// Mitsubishi GX Works2 project: 化成1_Debug 5.21   PLC: Q06UDEH

TYPE SwitchIO : STRUCT
  xLiftCylinderRetractDetect : BOOL;
  xLiftCylinderExtendDetect : BOOL;
  xLiftCylinderRetract : BOOL;
  xLiftCylinderExtend : BOOL;
  xEntryBarCylinderRetract : BOOL;
  xLiftCylinderExtendInit : BOOL;
  xEntryEnable : BOOL;
  xExitEnable : BOOL;
  xExitBarCylinderRetract : BOOL;
  xSwithEnable : BOOL;
  xLiftCylinderRetractButton : BOOL;
  xLiftCylinderExtendButton : BOOL;
  xEntryBarCylinderRetractButton : BOOL;
  xExitBarCylinderRetractButton : BOOL;
END_STRUCT END_TYPE

TYPE ConveyorIO : STRUCT
  iProductCategory : INT;  (* 产品类型0：无料1：正极  2：负极 3：隔膜 4：空料架 *)
  xCWPresent : BOOL;  (* 正转检测有无传感器 *)
  xCCWPresent : BOOL;  (* 反转检测有无传感器 *)
  xLoad : BOOL;  (* 上料请求 *)
  xUnload : BOOL;  (* 下料请求 *)
  xMotorCW : BOOL;  (* 电机正转 *)
  xMotorCCW : BOOL;  (* 电机反转 *)
  xEmpty : BOOL;  (* 线体状态为空 *)
  xNextRun : BOOL;  (* 下段线体运行 *)
  xUnloadCCW : BOOL;  (* 下料为反转 *)
  xloadCCW : BOOL;  (* 上料为反转 *)
  xLeave : BOOL;  (* 已经离开 *)
  xForward : BOOL;  (* 正转手动 *)
  xBackward : BOOL;  (* 反转手动 *)
  xBusy : BOOL;  (* 工作中 *)
  tLoadDelay : TIME;  (* 进入延时设置 *)
  xPutInto : BOOL;  (* 线体直接投入物料 *)
  xUnloadAlarm : BOOL;  (* 下料报警 *)
  xPosLimit : BOOL;  (* 正限位 *)
  xNegLimit : BOOL;  (* 负限位 *)
  xOverWidthAlarm : BOOL;  (* 超宽报警 *)
  xLimitAlarrm : BOOL;  (* 限位报警 *)
  iDeviceID : INT;  (* 线体ID *)
  xSizeDeficientDetect : BOOL;  (* 尺寸不足检测标志位 *)
END_STRUCT END_TYPE

TYPE ShuttleCarIO : STRUCT
  xReady : BOOL;  (* 准备就绪 *)
  xForward : BOOL;  (* 正转 *)
  xBackward : BOOL;  (* 反转 *)
  iCurrentPos : INT;  (* 当前位置 *)
  iDestinationPos : INT;  (* 目标位置 *)
  xCW : BOOL;  (* 正转输出 *)
  xCCW : BOOL;  (* 反转输出 *)
  xBrake : BOOL;  (* 刹车 *)
  xHomeSwitch : BOOL;  (* 零位接近开关 *)
  xPosLimit : BOOL;  (* 正限位 *)
  xNegLimit : BOOL;  (* 负限位 *)
  xMDIExe : BOOL;  (* MDI开始 *)
  xMDIDone : BOOL;  (* MDI 完成 *)
  xPassLimit : BOOL;  (* 限位屏蔽 *)
  xPosLimitCatch : BOOL;  (* 正限位捕捉 *)
  xNegLimitCatch : BOOL;  (* 负限位捕捉 *)
  xHomeExe : BOOL;  (* 开始寻零 *)
  xHomeDone : BOOL;  (* 寻零完成 *)
  xHomeBusy : BOOL;  (* 寻零中 *)
  xHomeFailed : BOOL;  (* 寻零失败 *)
  xBusy : BOOL;  (* 工作中 *)
  tArriveDelay : TIME;  (* 到位延时 *)
  xCylinder : BOOL;  (* 气缸控制 *)
  tBrakeDelay : TIME;  (* 抱闸延时 *)
  xPauseRamp : BOOL;  (* 暂停减速斜坡标志位 *)
  xPresentDetect1 : BOOL;  (* 物料有无检测1 *)
  xPresentDetect2 : BOOL;  (* 物料有无检测2 *)
  xOvertimeAlarm : BOOL;  (* 超时报警 *)
  tSetOverTime : TIME;  (* 设置超时时间 *)
  xLooseDetect : BOOL;  (* 松绳检测 *)
  xLooseAlarm : BOOL;  (* 松绳报警 *)
END_STRUCT END_TYPE

TYPE Stub : STRUCT
  xLoadRequest : BOOL;
  xLoadRequestAkn : BOOL;
  xUnloadRequest : BOOL;
  xUnloadRequestAkn : BOOL;
END_STRUCT END_TYPE

TYPE RGVCommunication : STRUCT
  xFullLoadRequest : BOOL;  (* 满框上料请求 *)
  xFullUnloadRequest : BOOL;  (* 满框下料请求 *)
  xEmptyLoadRequest : BOOL;  (* 空框上料请求 *)
  xEmptyUnloadRequest : BOOL;  (* 空框下料请求 *)
  xFullLoadRequestAkn : BOOL;  (* 满框上料请求确认 *)
  xFullUnloadRequestAkn : BOOL;  (* 满框下料请求确认 *)
  xEmptyLoadRequestAkn : BOOL;  (* 空框上料请求确认 *)
  xEmptyUnloadRequestAkn : BOOL;  (* 空框下料请求确认 *)
  xFullLoadComplete : BOOL;  (* 满框上料完成 *)
  xFullUnloadComplete : BOOL;  (* 满框下料完成 *)
  xEmptyLoadComplete : BOOL;  (* 空框上料完成 *)
  xEmptyUnloadComplete : BOOL;  (* 空框下料完成 *)
  xFullLoadCompleteAkn : BOOL;  (* 满框上料完成确认 *)
  xFullUnloadCompleteAkn : BOOL;  (* 满框下料完成确认 *)
  xEmptyLoadCompleteAkn : BOOL;  (* 空框上料完成确认 *)
  xEmptyUnloadCompleteAkn : BOOL;  (* 空框下料完成确认 *)
  xMdiExe : BOOL;  (* RGV 执行 *)
  xMdiDone : BOOL;  (* RGV 执行完成 *)
  iCurrentPostion : INT;  (* RGV当前位置 *)
  iDestinationPos : INT;  (* RGV目标位置 *)
  xEmpty1 : BOOL;
  xNextRun1 : BOOL;
  xEmpty2 : BOOL;
  xNextRun2 : BOOL;
  xLoad1 : BOOL;
  xUnload1 : BOOL;
  xLoad2 : BOOL;
  xUnload2 : BOOL;
  xCollisionAlarm : BOOL;  (* 干涉报警 *)
  xRemoteReset : BOOL;  (* 远程复位 *)
  xAuto : BOOL;  (* 自动 *)
END_STRUCT END_TYPE

TYPE BarCylinderIO : STRUCT
  xPresentSwitch : BOOL;  (* 行程开关 *)
  xBarCylinder : BOOL;  (* 阻挡气缸 *)
  xEmpty : BOOL;  (* 为空指示 *)
  xTransportMotorCW : BOOL;  (* 输送电机正转 *)
  xUnload : BOOL;  (* 下料 *)
  xBarCylinderButton : BOOL;  (* 阻挡气缸 *)
  xTransportMotorCWButton : BOOL;  (* 输送电机正转按钮 *)
  xLoad : BOOL;  (* 上料 *)
  xNextRun : BOOL;  (* 下位设备开始运行 *)
  xTransportMotorCCWButton : BOOL;  (* 输送电机反转按钮 *)
  xTransportMotorCCW : BOOL;  (* 输送电机反转 *)
  iProductCategory : INT;  (* 产品种类 *)
  tLoadDelay : TIME;  (* 上料延时 *)
  xBarCylinderSecondary : BOOL;  (* 阻挡第二个无料的气缸 *)
  xBarSecondaryButton : BOOL;  (* 阻挡第二个无料的气缸手动按钮 *)
  iDeviceID : INT;  (* 设备编号 *)
END_STRUCT END_TYPE

// global labels: Global1
VAR_GLOBAL
  g_xAuto AT M11 : BOOL;
  g_xManual : BOOL;
  g_xEStop AT X23 : BOOL;
  g_xReset AT X20 : BOOL;
  g_xStackLampRed AT Y120 : BOOL;
  g_xStackLampAmber AT Y121 : BOOL;
  g_xStackLampGreen AT Y122 : BOOL;
  g_xBuzzer AT Y123 : BOOL;
  g_xStop AT M2 : BOOL;
  g_xLocalAutoStart AT M1 : BOOL;
  g_xRemoteAutoStart AT M0 : BOOL;
  g_xRemoteAuto AT M10 : BOOL;
  g_iState AT D40 : INT;
  g_iLocalAutoStep : BOOL;
  g_xAlarm : BOOL;
  g_xImport1Forbidden AT M174 : BOOL;  (* 1表示禁止从注液入库 *)
  g_xExportChemForbidden AT M176 : BOOL;  (* 1表示禁止出库到化成 *)
  g_xExportBackForbidden AT M177 : BOOL;  (* 1表示禁止返回注液 *)
  g_xImport2Forbidden AT M175 : BOOL;  (* 1表示禁止从化成入库 *)
  g_xResetSingle AT M4 : BOOL;  (* 单线体复位 *)
  g_xInsertTask AT M5 : BOOL;  (* 插入任务 *)
  g_iInsertTask AT D2 : INT;  (* 插入任务号 *)
  g_xPause AT M3 : BOOL;  (* 暂停 *)
  g_iDeviceIDSelect AT D0 : INT;
END_VAR

// global labels: Global
VAR_GLOBAL
  g_xChem2ComFailed : BOOL;
  g_xFillingRGVComFailed : BOOL;
END_VAR

// task Task_01 (event TRUE, interval 0, priority 31): POU, Start, UDP

PROGRAM POU
VAR
  H3000Conveyor1 : Conveyor;
  H3000Conveyor1IO : ConveyorIO;
  H3000Conveyor2 : Conveyor;
  H3000Conveyor2IO : ConveyorIO;
  H3000Conveyor3 : Conveyor;
  H3000Conveyor3IO : ConveyorIO;
  H3000Conveyor4 : Conveyor;
  H3000Conveyor4IO : ConveyorIO;
  H3000Conveyor5 : Conveyor;
  H3000Conveyor5IO : ConveyorIO;
  H3000Conveyor6 : Conveyor;
  H3000Conveyor6IO : ConveyorIO;
  H3000Conveyor7 : Conveyor;
  H3000Conveyor7IO : ConveyorIO;
  H3000Conveyor8 : Conveyor;
  H3000Conveyor8IO : ConveyorIO;
  H3000Conveyor9 : Conveyor;
  H3000Conveyor9IO : ConveyorIO;
  H3000Conveyor10 : Conveyor;
  H3000Conveyor10IO : ConveyorIO;
  H3000ChemConveyor1 : Conveyor;
  H3000ChemConveyor1IO : ConveyorIO;
  H3000ChemConveyor2 : Conveyor;
  H3000ChemConveyor2IO : ConveyorIO;
  H3000ChemConveyor3 : Conveyor;
  H3000ChemConveyor3IO : ConveyorIO;
  Lifter1 : ShuttleCar;
  Lifter1IO : ShuttleCarIO;
  Conveyor1 : Conveyor;
  Conveyor1IO : ConveyorIO;
  Lifter2 : ShuttleCar;
  Lifter2IO : ShuttleCarIO;
  Conveyor2 : Conveyor;
  Conveyor2IO : ConveyorIO;
  H2200Conveyor1 : Conveyor;
  H2200Conveyor1IO : ConveyorIO;
  H2200Conveyor2 : Conveyor;
  H2200Conveyor2IO : ConveyorIO;
  H2200Conveyor3 : Conveyor;
  H2200Conveyor3IO : ConveyorIO;
  H2200Conveyor4 : Conveyor;
  H2200Conveyor4IO : ConveyorIO;
  H2200Conveyor5 : Conveyor;
  H2200Conveyor5IO : ConveyorIO;
  H2200Conveyor6 : Conveyor;
  H2200Conveyor6IO : ConveyorIO;
  H2200Conveyor7 : Conveyor;
  H2200Conveyor7IO : ConveyorIO;
  H2200Conveyor8 : Conveyor;
  H2200Conveyor8IO : ConveyorIO;
  H2200Conveyor9 : Conveyor;
  H2200Conveyor9IO : ConveyorIO;
  H2200Conveyor10 : Conveyor;
  H2200Conveyor10IO : ConveyorIO;
  H1000Conveyor1 : Conveyor;
  H1000Conveyor1IO : ConveyorIO;
  H1000Conveyor2 : Conveyor;
  H1000Conveyor2IO : ConveyorIO;
  H1000Conveyor3 : Conveyor;
  H1000Conveyor3IO : ConveyorIO;
  H1000Conveyor4 : Conveyor;
  H1000Conveyor4IO : ConveyorIO;
  H1000Conveyor5 : Conveyor;
  H1000Conveyor5IO : ConveyorIO;
  H1000Conveyor6 : Conveyor;
  H1000Conveyor6IO : ConveyorIO;
  H1000Conveyor7 : Conveyor;
  H1000Conveyor7IO : ConveyorIO;
  H1000Conveyor8 : Conveyor;
  H1000Conveyor8IO : ConveyorIO;
  H1000Conveyor9 : Conveyor;
  H1000Conveyor9IO : ConveyorIO;
  H3000SwitchChem : Switch;
  H3000SwitchChemIO : SwitchIO;
  H850Switch : Switch;
  H850SwitchIO : SwitchIO;
  H850SwitchConveyorIn : ConveyorIO;
  H850SwitchConveyorOut : ConveyorIO;
  H850Conveyor8 : Conveyor;
  H850Conveyor8IO : ConveyorIO;
  H1000Conveyor10 : Conveyor;
  H1000Conveyor10IO : ConveyorIO;
  H3000SwitchChemConveyorIn : ConveyorIO;
  H3000SwitchChemConveyorOut : ConveyorIO;
  H3000SwitchQuadPackage : Switch;
  H3000SwitchQuadPackageIO : SwitchIO;
  H3000SwitchPackageConveyorIn : ConveyorIO;
  H3000SwitchPackageConveyorOut : ConveyorIO;
  H2200Switch1 : Switch;
  H2200Switch1IO : SwitchIO;
  H2200Switch1ConveyorIn : ConveyorIO;
  H2200Switch1ConveyorOut : ConveyorIO;
  H2200Switch2 : Switch;
  H2200Switch2IO : SwitchIO;
  H2200Switch2ConveyorIn : ConveyorIO;
  H2200Switch2ConveyorOut : ConveyorIO;
  iStep : INT;
  Import1Conveyor1 : Conveyor;
  Import1Conveyor1IO : ConveyorIO;
  Import1Conveyor2 : Conveyor;
  Import1Conveyor2IO : ConveyorIO;
  Import2Conveyor1 : Conveyor;
  Import2Conveyor1IO : ConveyorIO;
  Import2Conveyor2 : Conveyor;
  Import2Conveyor2IO : ConveyorIO;
  Export1Conveyor1 : Conveyor;
  Export1Conveyor1IO : ConveyorIO;
  Export1Conveyor2 : Conveyor;
  Export1Conveyor2IO : ConveyorIO;
  Export2Conveyor1 : Conveyor;
  Export2Conveyor1IO : ConveyorIO;
  Export2Conveyor2 : Conveyor;
  Export2Conveyor2IO : ConveyorIO;
  Export2Switch : Switch;
  Export2SwitchIO : SwitchIO;
  Export2SwitchConveyorIn : ConveyorIO;
  Export2SwitchConveyorOut : ConveyorIO;
  H850Rotor : ShuttleCar;
  H850RotorIO : ShuttleCarIO;
  H850RotorConveyor : Conveyor;
  H850RotorConveyorIO : ConveyorIO;
  H2200RotorIO : ShuttleCarIO;
  H2200RotorConveyor : Conveyor;
  H2200RotorConveyorIO : ConveyorIO;
  H2200Rotor : ShuttleCar;
  H850Conveyor1 : Conveyor;
  H850Conveyor1IO : ConveyorIO;
  H850Conveyor3 : Conveyor;
  H850Conveyor3IO : ConveyorIO;
  H850Conveyor4 : Conveyor;
  H850Conveyor4IO : ConveyorIO;
  H850Conveyor5 : Conveyor;
  H850Conveyor5IO : ConveyorIO;
  H850Conveyor6 : Conveyor;
  H850Conveyor6IO : ConveyorIO;
  Lifter2Position : ARRAY [0..5] OF INT;
  ii : INT;  (* 提升机2任务号 *)
  H2200SwitchEmptyABack : Switch;
  H2200SwitchEmptyABackIO : SwitchIO;
  H2200SwitchEmptyABackConveyorIn : ConveyorIO;
  H2200SwitchEmptyABackConveyorOut : ConveyorIO;
  H2200SwitchEmptyBBack : Switch;
  H2200SwitchEmptyBBackIO : SwitchIO;
  H2200SwitchEmptyBBackConveyorIn : ConveyorIO;
  H2200SwitchEmptyBBackConveyorOut : ConveyorIO;
  H2200ImportConveyor1 : Conveyor;
  H2200ImportConveyor1IO : ConveyorIO;
  H2200ImportConveyor2 : Conveyor;
  H2200ImportConveyor2IO : ConveyorIO;
  Import1Switch : Switch;
  Import1SwitchIO : SwitchIO;
  Import1SwitchConveyorIn : ConveyorIO;
  Import1SwitchConveyorOut : ConveyorIO;
  Export1Switch : Switch;
  Export1SwitchIO : SwitchIO;
  Export1SwitchConveyorIn : ConveyorIO;
  Export1SwitchConveyorOut : ConveyorIO;
  Import2Switch : Switch;
  Import2SwitchIO : SwitchIO;
  Import2SwitchConveyorIn : ConveyorIO;
  Import2SwitchConveyorOut : ConveyorIO;
  Import1LoadCylinder : ShuttleCar;
  Import1LoadCylinderIO : ShuttleCarIO;
  Import2LoadCylinder : ShuttleCar;
  Import2LoadCylinderIO : ShuttleCarIO;
  Export1LoadCylinder : ShuttleCar;
  Export1LoadCylinderIO : ShuttleCarIO;
  Export2LoadCylinder : ShuttleCar;
  Export2LoadCylinderIO : ShuttleCarIO;
  Lifter2ExportChem : BOOL;  (* 提升机2满框去化成 *)
  Lifter2TaskID : INT;  (* 提升机2动作步骤 *)
  Lifter2Task : PriorityFB;
  H2200Switch1Task : PriorityFB;
  H2200Switch1TaskID : INT;
  H2200Switch1EmptyImport : BOOL;  (* 空框返回入库 *)
  Lifter1Speed : ShuttleCarVelocityFB;
  xScaning1 : BOOL;  (* 第1次扫码中，暂时停止运行 *)
  xScaning2 : BOOL;  (* 第2次扫码中，暂时停止运行 *)
  H850Conveyor7 : Conveyor;
  H850Conveyor7IO : ConveyorIO;
  H2200ImportConveyor3 : Conveyor;
  H2200ImportConveyor3IO : ConveyorIO;
  m_iExportConveyorOcuppy : INT;  (* 0:无占用1:1号出库 2:2号出库 *)
  m_tonExport2BayCylinderDalay : TON;
  m_xExport2BayCylinderDalay : BOOL;
  m_tExport2BayCylinderDalayCurren : TIME;
  m_tonImport1RequestDalay : TON;
  m_xImport1RequestDalay : BOOL;
  m_tImport1RequestDalaDalayCurren : TIME;
  m_tonImport2RequestDalay : TON;
  m_xImport2RequestDalay : BOOL;
  m_tImport2RequestDalaDalayCurren : TIME;
  m_tonHangUpChemDalay : TON;  (* 化成线阻塞延时 *)
  m_xHangUpChem : BOOL;  (* 化成线阻塞 *)
  m_tHangUpChemDalayCurrentTime : TIME;  (* 化成线阻塞 *)
  m_tonHangUpPackageDalay : TON;  (* 二封线阻塞 *)
  m_xHangUpPackage : BOOL;  (* 二封线阻塞 *)
  m_tHangUpPackageDalayCurrentTime : TIME;  (* 二封线阻塞当前时间 *)
  m_xImport2 : BOOL;  (* 出库线体使用间隔定时器 *)
  m_tonExportConveyorOcuppy : TON;  (* 出库线体使用间隔定时器 *)
  m_tExportConveyorOcuppyCurrent : TIME;
  m_xExportConveyorIdle : BOOL;  (* 出库线体空闲 *)
  m_tonScan2 : TON;  (* 扫码延时 *)
  m_tScan2 : TIME;  (* 扫码延时 *)
  m_xScan2 : BOOL;  (* 扫码延时 *)
  FillingStab1 : Stub;  (* 注液1号交互信号 *)
  FillingStab2 : Stub;  (* 注液2号交互信号 *)
  FillingStab3 : Stub;  (* 注液3号交互信号 *)
  FillingStab4 : Stub;  (* 注液4号交互信号 *)
  FillingRGV : RGVCommunication;
  H2200BayCylinderEmptyABack : BarCylinder;
  H2200BayCylinderEmptyABackIO : BarCylinderIO;
  H2200BayCylinderEmptyBBack : BarCylinder;
  H2200BayCylinderEmptyBBackIO : BarCylinderIO;
  m_xCartonARequest : BOOL;
  m_xCartonBRequest : BOOL;
  m_xCartonATaskLock : BOOL;
  m_xCartonBTaskLock : BOOL;
  m_xCartonALoadDone : BOOL;
  m_xCartonAStart : BOOL;
  m_xCartonBStart : BOOL;
  m_xCartonADone : BOOL;
  m_xCartonBDone : BOOL;
  FillQuarantineDoorInside : ShuttleCar;  (* 注液隔离门内部 *)
  FillQuarantineDoorInsideIO : ShuttleCarIO;  (* 注液隔离门内部 *)
  FillQuarantineDoorOutside : ShuttleCar;  (* 注液隔离门外部 *)
  FillQuarantineDoorOutsideIO : ShuttleCarIO;  (* 注液隔离门外部 *)
  m_xCartonADischargeLock : BOOL;  (* 下料锁，保证只下一个料框 *)
  m_xCartonBDischargeLock : BOOL;  (* 下料锁，保证只下一个料框 *)
  rejects1 : BOOL;  (* D线不良品 *)
  rejects2 : BOOL;  (* C线不良品 *)
  rejects3 : BOOL;  (* B线不良品 *)
  rejects4 : BOOL;  (* A线不良品 *)
  H850Conveyor2 : Conveyor;
  H850Conveyor2IO : ConveyorIO;
  ARorbidden : BOOL;  (* A线禁用 *)
  BRorbidden : BOOL;  (* B线禁用 *)
  CRorbidden : BOOL;  (* C线禁用 *)
  DRorbidden : BOOL;  (* D线禁用 *)
  TonScanAlarm1 : TON;
  TonScanAlarm2 : TON;
  TonScanAlarm3 : TON;
  TonScanAlarm1Time : TIME;
  TonScanAlarm2Time : TIME;
  TonScanAlarm3Time : TIME;
END_VAR
H3000SwitchQuadPackage(ConveyorEntryIO:=H3000SwitchPackageConveyorIn ,
                                                        ConveyorExitIO:=H3000SwitchPackageConveyorOut ,
                                                        SwitchIO:=H3000SwitchQuadPackageIO );
H3000SwitchQuadPackageIO.xLiftCylinderExtendButton:=M75;
H3000SwitchQuadPackageIO.xLiftCylinderRetractButton:=M76;
H3000SwitchQuadPackageIO.xExitBarCylinderRetractButton:=M83;
Y127:=H3000SwitchQuadPackageIO.xEXITBarCylinderRetract;
Y12C:=H3000SwitchQuadPackageIO.xLiftCylinderExtend;
Y12A:=H3000SwitchQuadPackageIO.xLiftCylinderRetract;
H3000SwitchQuadPackageIO.xLiftCylinderExtendDetect:=X29;
H3000SwitchQuadPackageIO.xLiftCylinderRetractDetect:=X2A;
H3000SwitchPackageConveyorIn.xForward:=M77;
H3000SwitchPackageConveyorIn.xCWPresent:=X28;
(*Y187:=H3000SwitchPackageConveyorIn.xMotorCW;*)
H3000SwitchPackageConveyorIn.iDeviceID:=3099;
H3000SwitchPackageConveyorOut.xForward:=M78;
H3000SwitchPackageConveyorOut.xCWPresent:=X2B;
Y12B:=H3000SwitchPackageConveyorOut.xMotorCW;
H3000SwitchPackageConveyorOut.iDeviceID:=3099;

H3000SwitchChem(ConveyorEntryIO:=H3000SwitchChemConveyorIn ,
                                                        ConveyorExitIO:=H3000SwitchChemConveyorOut ,
                                                        SwitchIO:=H3000SwitchChemIO );
H3000SwitchChemIO.xLiftCylinderExtendButton:=M79;
H3000SwitchChemIO.xLiftCylinderRetractButton:=M80;
Y129:=H3000SwitchChemIO.xLiftCylinderExtend;
Y12D:=H3000SwitchChemIO.xLiftCylinderRetract;
H3000SwitchChemIO.xLiftCylinderExtendDetect:=X2C;
H3000SwitchChemIO.xLiftCylinderRetractDetect:=X2D;
H3000SwitchChemConveyorIn.xForward:=M81;
H3000SwitchChemConveyorIn.xCWPresent:=X27;
H3000SwitchChemConveyorIn.tLoadDelay:=T#1s;
(*Y19B:=H3000SwitchPackageConveyorIn.xMotorCW;*)
H3000SwitchChemConveyorIn.iDeviceID:=3098;
H3000SwitchChemConveyorOut.xForward:=M82;
H3000SwitchChemConveyorOut.xCWPresent:=X2E;
Y12E:=H3000SwitchChemConveyorOut.xMotorCW;
H3000SwitchChemIO.xSwithEnable:=1;
H3000SwitchChemConveyorOut.iDeviceID:=3098;

Lifter1(ShuttleCarInOut:=Lifter1IO);
ShuttleCarCurrentPosition(X8C OR X8D ,X8C ,X8D, FALSE, Lifter1IO.iCurrentPos);
Lifter1Speed(xEnable:= g_xAuto,
                        xMotorCW:= Lifter1IO.xCW ,
                        xMotorCCW:= Lifter1IO.xCCW,
                        xPosition1Switch:= X8C,
                        xDecelerationSwitch:= X8B ,
	                    xPosition2Switch:= X8D ,
	                    xHighSpeed:= Y18F );
Lifter1IO.xReady:=X24;
Lifter1Io.xForward:=M50 OR X91;
Lifter1IO.xBackward:=M51 OR X92;
Lifter1IO.xPosLimit:=X8E;
Lifter1IO.xNegLimit:=X8F;
Y18D:=Lifter1IO.xCW;
Y18E:=Lifter1IO.xCCW;
Y192:=Lifter1IO.xBrake;

Conveyor1(ConveyorMotor:=Conveyor1IO);
Conveyor1IO.xForward:=M52;
Conveyor1IO.xBackward:=M53;
Conveyor1IO.xCWPresent:=X93;
Conveyor1IO.xCCWPresent:=X94;
Y18B:=Conveyor1IO.xMotorCW AND (X10B OR X8D) ;
Y18C:=Conveyor1IO.xMotorCCW AND X10B;
Conveyor1IO.xSizeDeficientDetect:=1;
Conveyor1IO.iDeviceID:=1;
(*2号提升机*)
Lifter2(ShuttleCarInOut:=Lifter2IO);
Lifter2Position[0]:=0;
Lifter2Position[1]:=128;
Lifter2Position[2]:=624;
Lifter2Position[3]:=5862;(*-----我改了一些位置，1层57•••77,4层6202•••6152*)
Lifter2Position[4]:=6178;
Lifter2Position[5]:=9230;
Y195:=ShuttleCarVelocityEncoder( g_xAuto , D190 , Lifter2Position[Lifter2IO.iDestinationPos] );
IF LDP(TRUE,g_xAuto) THEN
	Lifter2IO.iCurrentPos:=0;
END_IF;
FOR ii:=0 TO 5 BY 1 DO
	IF abs(D190-Lifter2Position[ii])<10 THEN
		Lifter2IO.iCurrentPos:=ii;
	END_IF;
END_FOR;
Lifter2IO.xReady:=X25;
(*提升机占用标志位控制*)(*-----这里我写了触摸屏M3、M4、M5、M6来控制各任务许可*)
Lifter2Task(xCondition1:= NOT H850Conveyor8IO.xEmpty AND  NOT g_xImport1Forbidden AND H2200ImportConveyor2IO.xEmpty AND D2340=2,
                     xCondition2:= NOT H1000Conveyor1IO.xEmpty AND NOT g_xImport2Forbidden AND H2200ImportConveyor2IO.xEmpty ,
                     xCondition3:= NOT H3000ChemConveyor3IO.xEmpty  AND (D2310=3 OR  D2310=2) AND NOT g_xExportChemForbidden AND H2200Conveyor1IO.xEmpty,
                     xCondition4:= NOT H3000ChemConveyor3IO.xEmpty  AND D2310=5 AND NOT g_xExportBackForbidden AND  H2200ImportConveyor2IO.xEmpty,
                     xCondition5:= FALSE ,(**)
	                 xTaskComplete:= (Lifter2IO.iCurrentPos=3 OR Lifter2IO.iCurrentPos=4) AND LDP(TRUE,Conveyor2IO.xEmpty)  ,
	                 xReset:= g_xReset,
	                 iPriority:=  Lifter2TaskID );
Lifter2Io.xForward:=M54 OR X9B;
Lifter2IO.xBackward:=M55 OR X9C;
Lifter2IO.xPosLimit:=X98;
Lifter2IO.xNegLimit:=X99;
Lifter2IO.xLooseDetect:=X9A;
Y193:=Lifter2IO.xCW;
Y194:=Lifter2IO.xCCW;
Y198:=Lifter2IO.xBrake;
(*提升机2编码器清零，到达负限位后清零*)
IF NOT Lifter2IO.xNegLimit THEN
	Y125:=1;
ELSE
	Y125:=0;
END_IF;

Conveyor2(ConveyorMotor:=Conveyor2IO);
Conveyor2IO.xForward:=M56;
Conveyor2IO.xBackward:=M57;
Conveyor2IO.xCWPresent:=X9D;
Conveyor2IO.xCCWPresent:=X9E;
Y19A:=Conveyor2IO.xMotorCW;
Y199:=Conveyor2IO.xMotorCCW;
Conveyor2IO.xSizeDeficientDetect:=1;(*不能增加尺寸检测，限位开关容易折断*)
Conveyor2IO.tLoadDelay:=T#200ms;
Conveyor2IO.iDeviceID:=2;
(*去二封线体*)
H3000Conveyor1(ConveyorMotor:=H3000Conveyor1IO);
H3000Conveyor1IO.xForward:=M30;
H3000Conveyor1IO.xCWPresent:=X2F;
Y12F:=H3000Conveyor1IO.xMotorCW;
H3000Conveyor1IO.iDeviceID:=3001;

H3000Conveyor2(ConveyorMotor:=H3000Conveyor2IO);
H3000Conveyor2IO.xForward:=M31;
H3000Conveyor2IO.xCWPresent:=X30;
Y130:=H3000Conveyor2IO.xMotorCW;
H3000Conveyor2IO.iDeviceID:=3002;

H3000Conveyor3(ConveyorMotor:=H3000Conveyor3IO);
H3000Conveyor3IO.xForward:=M32;
H3000Conveyor3IO.xCWPresent:=X31;
Y131:=H3000Conveyor3IO.xMotorCW;
H3000Conveyor3IO.iDeviceID:=3003;

H3000Conveyor4(ConveyorMotor:=H3000Conveyor4IO);
H3000Conveyor4IO.xForward:=M33;
H3000Conveyor4IO.xCWPresent:=X32;
Y132:=H3000Conveyor4IO.xMotorCW;
H3000Conveyor4IO.iDeviceID:=3004;

H3000Conveyor5(ConveyorMotor:=H3000Conveyor5IO);
H3000Conveyor5IO.xForward:=M34;
H3000Conveyor5IO.xCWPresent:=X33;
Y133:=H3000Conveyor5IO.xMotorCW;
H3000Conveyor5IO.iDeviceID:=3005;

H3000Conveyor6(ConveyorMotor:=H3000Conveyor6IO);
H3000Conveyor6IO.xForward:=M34;
H3000Conveyor6IO.xCWPresent:=X34;
Y134:=H3000Conveyor6IO.xMotorCW;
H3000Conveyor6IO.iDeviceID:=3006;

H3000Conveyor7(ConveyorMotor:=H3000Conveyor7IO);
H3000Conveyor7IO.xForward:=M35;
H3000Conveyor7IO.xCWPresent:=X35;
Y135:=H3000Conveyor7IO.xMotorCW;
H3000Conveyor7IO.iDeviceID:=3007;

H3000Conveyor8(ConveyorMotor:=H3000Conveyor8IO);
H3000Conveyor8IO.xForward:=M36;
H3000Conveyor8IO.xCWPresent:=X36;
Y136:=H3000Conveyor8IO.xMotorCW;
H3000Conveyor8IO.iDeviceID:=3008;

H3000Conveyor9(ConveyorMotor:=H3000Conveyor9IO);
H3000Conveyor9IO.xForward:=M37;
H3000Conveyor9IO.xCWPresent:=X37;
Y137:=H3000Conveyor9IO.xMotorCW;
H3000Conveyor9IO.iDeviceID:=3009;

H3000Conveyor10(ConveyorMotor:=H3000Conveyor10IO);
H3000Conveyor10IO.xForward:=M38;
H3000Conveyor10IO.xCWPresent:=X38;
Y138:=H3000Conveyor10IO.xMotorCW;
H3000Conveyor10IO.iDeviceID:=3010;

(*本段线体没有接线*)
(*H3000ChemConveyor1(ConveyorMotor:=H3000ChemConveyor1IO);
H3000ChemConveyor1IO.xForward:=M39;
H3000ChemConveyor1IO.xCWPresent:=X39;
Y139:=H3000ChemConveyor1IO.xMotorCW;*)

(*去化成H3000线体*)
H3000ChemConveyor2(ConveyorMotor:=H3000ChemConveyor2IO);
H3000ChemConveyor2IO.xForward:=M40;
H3000ChemConveyor2IO.xCWPresent:=X39;
Y13A:=H3000ChemConveyor2IO.xMotorCW;
H3000ChemConveyor2IO.iDeviceID:=3092;

H3000ChemConveyor3(ConveyorMotor:=H3000ChemConveyor3IO);
H3000ChemConveyor3IO.xForward:=M41;
H3000ChemConveyor3IO.xCWPresent:=X3B;
H3000ChemConveyor3IO.xPosLimit:=NOT X3A;
Y13B:=H3000ChemConveyor3IO.xMotorCW;
H3000ChemConveyor3IO.iDeviceID:=3093;
(*入库线体*)
H2200Switch1(ConveyorEntryIO:=H2200Switch1ConveyorIn ,
                                                        ConveyorExitIO:=H2200Switch1ConveyorOut ,
                                                        SwitchIO:=H2200Switch1IO );
m_xCartonARequest:=XAE OR XAA OR XA6  ;
m_xCartonBRequest:=XA2;
 IF  m_xCartonARequest  (*A空框上料请求信号*)
 	AND NOT m_xCartonAStart 
 	AND  NOT m_xCartonBStart 
 	AND H2200Switch1TaskID<>1  THEN
 	 m_xCartonAStart:=1;
 	 m_xCartonATaskLock:=1;(*任务锁，保证一次呼叫只执行一次出空框任务*)
 END_IF;   
 IF  H2200Switch1TaskID=1 THEN
 	m_xCartonATaskLock:=0;
 END_IF; 
  IF  m_xCartonBRequest  (*B空框上料请求信号*)
  	AND  NOT m_xCartonBStart 
  	AND NOT m_xCartonAStart 
  	AND H2200Switch1TaskID<>2   THEN
 	 m_xCartonBStart:=1;
 	 m_xCartonBTaskLock:=1;(*任务锁，保证一次呼叫只执行一次出空框任务*)
  END_IF;
  IF H2200Switch1TaskID=2 THEN
  	m_xCartonBTaskLock:=0;
  END_IF;
  IF m_xCartonADone OR g_xReset OR g_xManual OR LDF(TRUE,H850Conveyor1IO.xEmpty) THEN                                               
		m_xCartonAStart:=0;
  END_IF;
   IF m_xCartonBDone OR g_xReset OR g_xManual OR LDF(TRUE,H850Conveyor1IO.xEmpty) THEN                                               
		m_xCartonBStart:=0;
   END_IF; 
H2200Switch1Task(xCondition1:=H2200SwitchEmptyABackConveyorIn.xEmpty   (*倍速链前顶升移载为空*)
															AND NOT H2200Switch1EmptyImport                  (*无入库*)
															AND NOT H2200BayCylinderEmptyABackIO.xEmpty (*倍速链有料*)
															AND H2200RotorConveyorIO.xEmpty(*转台为空*)
															AND NOT H2200RotorConveyorIO.xBusy,(*转台无工作中信号*)
															(*AND m_xCartonATaskLock,(*任务锁*)
                                    xCondition2:=H2200SwitchEmptyBBackConveyorIn.xEmpty   (*倍速链前顶升移载为空*)
                                    						AND NOT H2200Switch1EmptyImport                  (*无入库*)
                                    						AND NOT H2200BayCylinderEmptyBBackIO.xEmpty (*倍速链有料*)
                                    						AND H2200RotorConveyorIO.xEmpty(*转台为空*)
                                    						AND NOT H2200RotorConveyorIO.xBusy ,
                                    						(*AND m_xCartonBTaskLock,(*任务锁*)
                                    xCondition3:=(*NOT  H2200SwitchEmptyABackConveyorIn.xEmpty AND NOT H2200Switch1EmptyImport AND X5D*) FALSE  ,
                                    xCondition4:=(* NOT  H2200SwitchEmptyBBackConveyorIn.xEmpty AND NOT H2200Switch1EmptyImport and x4c*)FALSE,
                                    xCondition5:= NOT H2200ImportConveyor3IO.xEmpty AND H2200ImportConveyor1IO.xEmpty ,
	                               xTaskComplete:= LDP(TRUE, H2200Switch1ConveyorIn.xEmpty) OR LDP(TRUE, H2200Switch1ConveyorOut.xEmpty)  ,
	                               xReset:= g_xResetSingle AND g_iDeviceIDSelect=2299 ,
	                               iPriority:= H2200Switch1TaskID);
H2200Switch1IO.xLiftCylinderExtendButton:=M84;
H2200Switch1IO.xLiftCylinderRetractButton:=M85;
H2200Switch1IO.xExitBarCylinderRetractButton:=M86;
Y158:=H2200Switch1IO.xEXITBarCylinderRetract;
Y155:=H2200Switch1IO.xLiftCylinderExtend;
Y156:=H2200Switch1IO.xLiftCylinderRetract;
H2200Switch1IO.xLiftCylinderExtendDetect:=X55;
H2200Switch1IO.xLiftCylinderRetractDetect:=X56;
H2200Switch1ConveyorIn.xForward:=M87;
H2200Switch1ConveyorIn.xCWPresent:=X101;
H2200Switch1ConveyorIn.iDeviceID:=2299;
H2200Switch1ConveyorIn.tLoadDelay:=T#5s;
(*Y177:=H2200Switch1ConveyorIn.xMotorCW;*)
H2200Switch1ConveyorOut .xForward:=M88;
H2200Switch1ConveyorOut .xCWPresent:=X101;
H2200Switch1ConveyorOut.tLoadDelay:=T#1s;
Y157:=H2200Switch1ConveyorOut .xMotorCW;
H2200Switch1ConveyorOut .iDeviceID:=2299;

H2200ImportConveyor1(ConveyorMotor:=H2200ImportConveyor1IO);
H2200ImportConveyor1IO.xForward:=M136;
H2200ImportConveyor1IO.xCWPresent:=X53;
Y153:=H2200ImportConveyor1IO.xMotorCW;
H2200ImportConveyor1IO.iDeviceID:=2293;

H2200ImportConveyor2(ConveyorMotor:=H2200ImportConveyor2IO);
H2200ImportConveyor2IO.xForward:=M122;
H2200ImportConveyor2IO.xCWPresent:=X54;(*-----这里改了，X58•••X54*)
Y154:=H2200ImportConveyor2IO.xMotorCW;
H2200ImportConveyor2IO.iDeviceID:=2292;

H2200ImportConveyor3(ConveyorMotor:=H2200ImportConveyor3IO);
H2200ImportConveyor3IO.xForward:=M166;
H2200ImportConveyor3IO.xCWPresent:=X58;(*-----这里改了，X58•••X54*)
Y180:=H2200ImportConveyor3IO.xMotorCW;
H2200ImportConveyor3IO.iDeviceID:=2291;

H2200Switch2(ConveyorEntryIO:=H2200Switch2ConveyorIn ,
                                                        ConveyorExitIO:=H2200Switch2ConveyorOut ,
                                                        SwitchIO:=H2200Switch2IO );
H2200Switch2IO.xLiftCylinderExtendButton:=M89;
H2200Switch2IO.xLiftCylinderRetractButton:=M90;
H2200Switch2IO.xExitBarCylinderRetractButton:=M91;
Y15C:=H2200Switch2IO.xEXITBarCylinderRetract;
Y159:=H2200Switch2IO.xLiftCylinderExtend;
Y15A:=H2200Switch2IO.xLiftCylinderRetract;
H2200Switch2IO.xLiftCylinderExtendDetect:=X59;
H2200Switch2IO.xLiftCylinderRetractDetect:=X5A;
H2200Switch2ConveyorIn.xForward:=M92;
H2200Switch2ConveyorIn.xCWPresent:=X5B;
H2200Switch2ConveyorIn.tLoadDelay:=T#4s;
Y15B:=H2200Switch2ConveyorIn.xMotorCW;
H2200Switch2ConveyorIn.iDeviceID:=2298;
H2200Switch2ConveyorOut .xForward:=M93;
H2200Switch2ConveyorOut .xCWPresent:=X5B;
Y186:=H2200Switch2ConveyorOut.xMotorCW AND NOT xScaning1 ;(*	Y186:=1;(***入库倍速链***)(*-----这里加了xScaning扫码中*)
Y13C:=H2200Switch2ConveyorOut.xMotorCW AND NOT xScaning1 ;
Y19C:=H2200Switch2ConveyorOut.xMotorCW AND NOT xScaning1 ;
Y19D:=H2200Switch2ConveyorOut.xMotorCW AND NOT xScaning1 ;
H2200Switch2IO.xLiftCylinderExtendInit:=1;
H2200Switch2ConveyorOut.iDeviceID:=2298;

H2200BayCylinderEmptyABack(BarCylinderIO:= H2200BayCylinderEmptyABackIO );
H2200BayCylinderEmptyABackIO.xBarCylinderButton:=M189;
H2200BayCylinderEmptyABackIO.xPresentSwitch:=X5D;
Y15D:=H2200BayCylinderEmptyABackIO.xBarCylinder;
Y169:=H2200BayCylinderEmptyABackIO.xBarCylinderSecondary;

H2200BayCylinderEmptyBBack(BarCylinderIO:= H2200BayCylinderEmptyBBackIO);
H2200BayCylinderEmptyBBackIO.xBarCylinderButton:=M190;
H2200BayCylinderEmptyBBackIO.xPresentSwitch:=X6C;
Y16C:=H2200BayCylinderEmptyBBackIO.xBarCylinder;
Y16B:=H2200BayCylinderEmptyBBackIO.xBarCylinderSecondary;

H2200SwitchEmptyABack(ConveyorEntryIO:=H2200SwitchEmptyABackConveyorIn ,
                                                        ConveyorExitIO:=H2200SwitchEmptyABackConveyorOut ,
                                                        SwitchIO:=H2200SwitchEmptyABackIO );
H2200SwitchEmptyABackIO.xLiftCylinderExtendButton:=M137;
H2200SwitchEmptyABackIO.xLiftCylinderRetractButton:=M138;
H2200SwitchEmptyABackIO.xExitBarCylinderRetractButton:=M139;
Y160:=H2200SwitchEmptyABackIO.xLiftCylinderExtend;
Y161:=H2200SwitchEmptyABackIO.xLiftCylinderRetract;
H2200SwitchEmptyABackIO.xLiftCylinderExtendDetect:=X60;
H2200SwitchEmptyABackIO.xLiftCylinderRetractDetect:=X61;
H2200SwitchEmptyABackConveyorIn.xForward:=M140;
H2200SwitchEmptyABackConveyorIn.xCWPresent:=X62;
H2200SwitchEmptyABackConveyorIn.tLoadDelay:=T#2s;
Y162:=H2200SwitchEmptyABackConveyorIn.xMotorCW;
H2200SwitchEmptyABackConveyorIn.iDeviceID:=2295;
H2200SwitchEmptyABackConveyorOut .xForward:=M146;
H2200SwitchEmptyABackConveyorOut.xCWPresent:=X62;
H2200SwitchEmptyABackConveyorOut.iDeviceID:=2295;
(*空框返回共同倍速链*)
Y177:=H2200SwitchEmptyABackConveyorOut .xMotorCW 
			OR H2200SwitchEmptyBBackConveyorOut .xMotorCW 
			OR H2200Switch1ConveyorIn.xMotorCW;
Y181:=H2200SwitchEmptyABackConveyorOut .xMotorCW 
			OR H2200SwitchEmptyBBackConveyorOut .xMotorCW 
			OR H2200Switch1ConveyorIn.xMotorCW;

H2200SwitchEmptyBBack(ConveyorEntryIO:=H2200SwitchEmptyBBackConveyorIn ,
                                                        ConveyorExitIO:=H2200SwitchEmptyBBackConveyorOut ,
                                                        SwitchIO:=H2200SwitchEmptyBBackIO );
H2200SwitchEmptyBBackIO.xLiftCylinderExtendButton:=M141;
H2200SwitchEmptyBBackIO.xLiftCylinderRetractButton:=M142;
H2200SwitchEmptyBBackIO.xExitBarCylinderRetractButton:=M143;
Y166:=H2200SwitchEmptyBBackIO.xLiftCylinderExtend;
Y167:=H2200SwitchEmptyBBackIO.xLiftCylinderRetract;
H2200SwitchEmptyBBackIO.xLiftCylinderExtendDetect:=X66;
H2200SwitchEmptyBBackIO.xLiftCylinderRetractDetect:=X67;
H2200SwitchEmptyBBackConveyorIn.xForward:=M144;
H2200SwitchEmptyBBackConveyorIn.xCWPresent:=X68;
H2200SwitchEmptyBBackConveyorIn.tLoadDelay:=T#2s;
H2200SwitchEmptyBBackConveyorIn.iDeviceID:=2294;
Y168:=H2200SwitchEmptyBBackConveyorIn.xMotorCW;
H2200SwitchEmptyBBackConveyorOut .xForward:=M145;
H2200SwitchEmptyBBackConveyorOut.xCWPresent:=X68;
H2200SwitchEmptyBBackConveyorOut.iDeviceID:=2294;

(*空框回注液转台*)
H2200Rotor(ShuttleCarInOut:=H2200RotorIO);
ShuttleCarCurrentPosition(X6F OR X75 ,X75 ,X6F, FALSE,H2200RotorIO.iCurrentPos );
H2200RotorIO.xReady:=TRUE;
H2200RotorIO.xForward:=M78;
H2200RotorIO.xBackward:=M79;
H2200RotorIO.xPosLimit:=X72;
H2200RotorIO.xNegLimit:=X71;
Y170:=H2200RotorIO.xCW;
Y16F:=H2200RotorIO.xCCW;
Y1B8:=H2200RotorIO.xBrake;

H2200RotorConveyor(ConveyorMotor:=H2200RotorConveyorIO);
H2200RotorConveyorIO.xForward:=M80;
H2200RotorConveyorIO.xBackward:=M81;
H2200RotorConveyorIO.xCWPresent:=X74;
H2200RotorConveyorIO.xCcWPresent:=X73;
Y172:=H2200RotorConveyorIO.xMotorCW;
Y171:=H2200RotorConveyorIO.xMotorCCW;
H2200RotorConveyorIO.iDeviceID:=2280;
(*去化成H2200线体*)
H2200Conveyor1(ConveyorMotor:=H2200Conveyor1IO);
H2200Conveyor1IO.xForward:=M42;
H2200Conveyor1IO.xCWPresent:=X3F;
Y13F:=H2200Conveyor1IO.xMotorCW;
H2200Conveyor1IO.iDeviceID:=2201;

H2200Conveyor2(ConveyorMotor:=H2200Conveyor2IO);
H2200Conveyor2IO.xForward:=M43;
H2200Conveyor2IO.xCWPresent:=X40;
Y140:=H2200Conveyor2IO.xMotorCW;
H2200Conveyor2IO.iDeviceID:=2202;

H2200Conveyor3(ConveyorMotor:=H2200Conveyor3IO);
H2200Conveyor3IO.xForward:=M44;
H2200Conveyor3IO.xCWPresent:=X41;
Y141:=H2200Conveyor3IO.xMotorCW;
H2200Conveyor3IO.iDeviceID:=2203;

H2200Conveyor4(ConveyorMotor:=H2200Conveyor4IO);
H2200Conveyor4IO.xForward:=M45;
H2200Conveyor4IO.xCWPresent:=X42;
Y142:=H2200Conveyor4IO.xMotorCW;
H2200Conveyor4IO.iDeviceID:=2204;

H2200Conveyor5(ConveyorMotor:=H2200Conveyor5IO);
H2200Conveyor5IO.xForward:=M46;
H2200Conveyor5IO.xCWPresent:=X43;
Y143:=H2200Conveyor5IO.xMotorCW;
H2200Conveyor5IO.iDeviceID:=2205;

H2200Conveyor6(ConveyorMotor:=H2200Conveyor6IO);
H2200Conveyor6IO.xForward:=M47;
H2200Conveyor6IO.xCWPresent:=X44;
Y144:=H2200Conveyor6IO.xMotorCW;
H2200Conveyor6IO.iDeviceID:=2206;

H2200Conveyor7(ConveyorMotor:=H2200Conveyor7IO);
H2200Conveyor7IO.xForward:=M48;
H2200Conveyor7IO.xCWPresent:=X45;
Y145:=H2200Conveyor7IO.xMotorCW;
H2200Conveyor7IO.iDeviceID:=2207;

H2200Conveyor8(ConveyorMotor:=H2200Conveyor8IO);
H2200Conveyor8IO.xForward:=M49;
H2200Conveyor8IO.xCWPresent:=X46;
Y146:=H2200Conveyor8IO.xMotorCW;
H2200Conveyor8IO.iDeviceID:=2208;

H2200Conveyor9(ConveyorMotor:=H2200Conveyor9IO);
H2200Conveyor9IO.xForward:=M58;
H2200Conveyor9IO.xCWPresent:=X47;
Y147:=H2200Conveyor9IO.xMotorCW;
H2200Conveyor9IO.iDeviceID:=2209;

H2200Conveyor10(ConveyorMotor:=H2200Conveyor10IO);
H2200Conveyor10IO.xForward:=M59;
H2200Conveyor10IO.xCWPresent:=X48;
Y148:=H2200Conveyor10IO.xMotorCW;
H2200Conveyor10IO.iDeviceID:=2210;
(*去化成回流H1100线体*)
H1000Conveyor1(ConveyorMotor:=H1000Conveyor1IO);
H1000Conveyor1IO.xForward:=M60;
H1000Conveyor1IO.xCWPresent:=XDD;
H1000Conveyor1IO.xPosLimit:=NOT X49;
Y149:=H1000Conveyor1IO.xMotorCW;
H1000Conveyor1IO.iDeviceID:=1001;

H1000Conveyor2(ConveyorMotor:=H1000Conveyor2IO);
H1000Conveyor2IO.xForward:=M61;
H1000Conveyor2IO.xCWPresent:=X4A;
Y14A:=H1000Conveyor2IO.xMotorCW;
H1000Conveyor2IO.iDeviceID:=1002;

H1000Conveyor3(ConveyorMotor:=H1000Conveyor3IO);
H1000Conveyor3IO.xForward:=M62;
H1000Conveyor3IO.xCWPresent:=X4B;
Y14B:=H1000Conveyor3IO.xMotorCW;
H1000Conveyor3IO.iDeviceID:=1003;